// TIA Portal project "1215C_BREAKOUT_BOARD_IO-LINK_TEMPERATURE" (V19) (continued)
REGION Network 4: Add leading zero to HH:MM if less than 10
   // > If DTL.HOUR is less than 10 - replace 1st character in HH with a 0
   // > If DTL.MINUTE is less than 10 - replace 1st character in MM with a 0
   IF #LOCAL_DTL.HOUR < 10 THEN
       #sCustomTime_HH := REPLACE(IN1 := #sCustomTime_HH, IN2 := '0', L := 1, P := 1);
   END_IF;
   IF #LOCAL_DTL.MINUTE < 10 THEN
       #sCustomTime_MM := REPLACE(IN1 := #sCustomTime_MM, IN2 := '0', L := 1, P := 1);
   END_IF;
END_REGION

REGION Network 5: =================CONCAT_INTO_FORMAT=================
END_REGION

REGION Network 6: CONCAT Date into DD/MM/YY
   #sTemp_String := CONCAT(IN1 := #sCustomDate_DD, IN2 := '/');
   #sTemp_String := CONCAT(IN1 := #sTemp_String, IN2 := #sCustomDate_MM);
   #sTemp_String := CONCAT(IN1 := #sTemp_String, IN2 := '/');
   #sCustomDate_DDMMYY := CONCAT(IN1 := #sTemp_String, IN2 := #sCustomDate_YY);
END_REGION

REGION Network 7: CONCAT Time HH:MM
   #sCustomTime_HHMM := CONCAT(IN1 := #sCustomTime_HH, IN2 := ':');
   #sCustomTime_HHMM := CONCAT(IN1 := #sCustomTime_HHMM, IN2 := #sCustomTime_MM);
END_REGION
END_FUNCTION

// folder: WS01_TVET_Workstation/02-IOLink_Control

FUNCTION "FC10111-IFM_2Byte_PD" : Void   // FC10111, SCL
TITLE = IFM 2 Byte Process Data FC
{ S7_Optimized_Access := 'TRUE' }
VERSION : 0.1
// This function block is for a device with two byte process data input and no switch point in the 
// process data stream.
   VAR_INPUT
      I_PV : Int;   // input process value from master
      Gradient : Real;   // gradient see IODD descrption
   END_VAR
   VAR_OUTPUT
      O_PV_C : Real;   // output process value in deg c
      O_PV_F : Real;   // output process value in deg f
   END_VAR
   VAR_TEMP
      Temp_PV_C : Real;   // temp process value in deg c
   END_VAR
BEGIN
   // Convert input value using the gradient (default = 0.1)
   IF #Gradient > 0 THEN
       #Temp_PV_C := INT_TO_REAL(#I_PV) * #Gradient;
   ELSE
       #O_PV_C := INT_TO_REAL(#I_PV) * 1.0;
   END_IF;

   // Convert C to F
   #O_PV_F := (#Temp_PV_C * 1.8) + 32;

   // Move Temp_PV_C to O_PV_C
   #O_PV_C := #Temp_PV_C;
END_FUNCTION

// ===== library types =====

// folder: S7-1200/1500/Lib/S7-1200/1500/Common

FUNCTION_BLOCK "IO_LINK_DEVICE"   // FB50001, SCL
TITLE = IO_LINK_DEVICE
{ S7_Optimized_Access := 'TRUE' }
AUTHOR : SUP_FA
FAMILY : IO-Link
VERSION : 3.0
// Function block to read and write acyclic data on devices with IO-Link used on SIMATIC S7 controllers. (former IO_LINK_CALL)
   VAR_INPUT
      REQ : Bool;   // request function / Request Function / Neuer Auftrag
      ID : HW_IO;   // hardware identifier of IO-Link master module (HW_IO) from hw-config / Hardwarekennung des IOL-Master Moduls (HW_IO) aus HW-Konfiguration
      CAP : DInt := DINT#0;   // Client Access Point (CAP), for ET200 always 227 decimal / Client Access Point (CAP), bei ET200 immer 227 dez
      RD_WR : Bool;   // read and write access on IO-Link device 0: read, 1: write / Lese und Schreibzugriff auf IO-Link Device 0: Lesen, 1: schreiben
      PORT : Int := INT#0;   // number of port on IO-Link master module (ET200SP = 0..4) / Port/ Kanalnummer an dem das IO-Link Device betrieben wird. (ET200 = 0 .. 4)
      IOL_INDEX : Int := INT#0;   // address parameter Index (IO-Link Device) 0..32767 IOL-D, 65535 port functions / Adressparameter Index (IO-Link Device) 0..32767 IOL-D, 65535 port functions
      IOL_SUBINDEX : Int := INT#0;   // address parameter Subindex (IO-Link Device) 0 full record; 1-255 single parameter / Adressparameter Subindex (IO-Link Device) 0 ges. Record; 1-255 einz. Parameter
      LEN : Int := INT#0;   // length of writing data (netto data) / Länge der zu schreibenden Daten (Nettodaten)
   END_VAR
   VAR_OUTPUT
      DONE_VALID : Bool;   // validity 0: data invalid ; 1: data valid / Gültigkeit 0: Daten nicht gültig; 1: Daten gültig
      BUSY : Bool;   // 0: request finish 1: request in progress / 0: Auftrag abgeschlossen 1: Auftrag in Bearbeitung
      ERROR : Bool;   // Error Flag = 0: no error; 1: function aborted with error / Fehler Flag 0: kein Fehler; 1: Abbruch der Funktion mit Fehler
      STATUS : DWord := DW#16#00000000;   // DP/ PNIO - error status ; ERROR Flag = 1 - communication error status in detail / DP/ PNIO - Fehlerstatus; ERROR Flag = 1 - detaillierter Kommunikationsfehlerstatus
      IOL_STATUS : DWord := DW#16#00000000;   // IO-Link error status; ERROR flag = 1: IO-Link error status in detail / IO-Link Fehlerstatus; ERROR Flag = 1 - detaillierte IO-Link Fehlerstatus
      RD_LEN : Int := INT#0;   // length of read data record (number of bytes) / Länge des gelesenen Datensatzes (Anzahl Bytes)
   END_VAR
   VAR_IN_OUT
      RECORD_IOL_DATA : Array[0..231] of Byte;   // data area for reading / writing data (max. 232 byte) / Datenbereich für LESEN / SCHREIBEN (max. 232 Byte)
   END_VAR
   VAR
      RDREC_Function : RDREC;   // system function "read data record" (former SFB52) / Funktion Datensatz lesen (ehemals SFB52)
      WRREC_Function : WRREC;   // system function "write data record" (former SFB53) / Funktion Datensatz schreiben (ehemals SFB53)
      TP_poll : TP_TIME;   // poll rate read data record / Pollzeit für "Datensatz lesen"
      TON_monitoring : TON_TIME;   // request monitoring time / Überwachungszeit für Aufträge
      rdrec : Struct   // internal structure for RDREC / interne Struktur für RDREC
         valid : Bool;   // Function performed
         busy : Bool;   // Function busy
         error : Bool;   // Error flag
         status : DWord;   // Function result/error message
         length : UInt;   // Length of the fetched data record
      END_STRUCT;
      wrrec : Struct   // internal structure for WRREC / interne Struktur für WRREC
         length : UInt;   // length of write data record
         done : Bool;   // Function performed
         busy : Bool;   // Function busy
         error : Bool;   // Error flag
         status : DWord;   // Function result/error message
      END_STRUCT;
      read : Struct   // data area for reading data / Datenbereich für Lesedaten
         header : Struct
            CALL : Struct   // header for read/write data record
               Extended_Function_Num : Byte := 16#8;   // extended function number (fix coded 08h)
               Port : Byte;   // variable port (user interface) 0...255
               FI_Index : Word := 16#FE4A;   // FI index (fix coded 65098)
            END_STRUCT;
            IOL : Struct   // header for IO-Link
               Control : Byte;   // RD_WR = 0 = read = Control:=0x03 / / RD_WR = 1 = write = Control:=0x02
               Index_HighByte : Byte;   // index of data record 0…32767 (high byte)
               Index_LowByte : Byte;   // index of data record 0…32767 (low byte)
               Subindex : Byte;   // subindex for data record 0...255
            END_STRUCT;
         END_STRUCT;
         data : Array[0..231] of Byte;
      END_STRUCT;
      write : Struct   // data area for writing data / Datenbereich für Schreibdaten
         header : Struct
            CALL : Struct   // header for read/write data record
               Extended_Function_Num : Byte := 16#8;   // extended function number (fix coded 08h)
               Port : Byte;   // variable port (user interface) 0...255
               FI_Index : Word := 16#FE4A;   // FI index (fix coded 65098)
            END_STRUCT;
            IOL : Struct   // header for IO-Link
               Control : Byte;   // RD_WR = 0 = read = Control:=0x03 / / RD_WR = 1 = write = Control:=0x02
               Index_HighByte : Byte;   // index of data record 0…32767 (high byte)
               Index_LowByte : Byte;   // index of data record 0…32767 (low byte)
               Subindex : Byte;   // subindex for data record 0...255
            END_STRUCT;
         END_STRUCT;
         data : Array[0..231] of Byte;
      END_STRUCT;
      sequencecontrol : Int := INT#0;   // number of sequence control
      typeofrequest : Int := INT#0;   // type of request (0=Read, 1=Write)
      R_TRIG_REQ : Bool;   // impulse start new request / Impuls für neuen Auftrag starten
      R_TRIG_REQ_old : Bool;   // old value of REQ (previous cycle) / Flankenmerker
      F_TRIG_poll : Bool;   // impulse poll read data record (response) / Impuls für Pollen "Datensatz lesen"
      F_TRIG_poll_old : Bool;   // old value of Poll (previous cycle) / Flankenmerker
   END_VAR
   VAR_TEMP
      retval : Int;   // function return value / Variable für Rückgabewerte von Funktionen
      tmpWORD : Word;   // data type WORD for temporarily use / Datentyp WORD zur temporären Verwendung
      tmpDWORD : DWord;   // data type DWORD for temporarily use / Datentyp DWORD zur temporären Verwendung
      tmpINT : Int;   // data type INT for temporarily use / Datentyp INT zur temporären Verwendung
      i : Int;   // run tag for counting loops / Laufvariable für for-Schleifen
   END_VAR
BEGIN
   (*---------------------------------------------------------------------------------------------------------------------
   SIEMENS AG
   ©Copyright 2015. All Rights Reserved.
   -----------------------------------------------------------------------------------------------------------------------
   Limitation of liability
   This software was developed with largest care. However, the author can not guarantee, that the software runs under
   each version of STEP7 on each PLC flawlessly.
   There is no warranty for the software, to the extent permitted by applicable law. The copyright holder provides the
   software "as is" without warranty of any kind, either expressed or implied, including, but not limited to, the implied
   warranties of merchantability and fitness for a particular purpose. The entire risk as to the quality and performance
   of the software is with you. Should the software prove defective, you assume the cost of all necessary servicing,
   repair or correction. In no event unless required by applicable law will the copyright holder be liable to you for
   damages, including any general, special, incidental or consequential damages arising out of the use or inability to
   use the software (including but not limited to loss of data or data being rendered inaccurate or losses sustained by
   you or third parties or a failure of the software to operate with any other programs), even if such holder or other
   party has been advised of the possibility of such damages.
   Permission to use or copy this software for any purpose is hereby granted without fee, provided the above notices are
   retained on all copies. Permission to modify the code and to distribute modified code is granted, provided the above
   notices are retained, and a notice that the code was modified is included with the above copyright notice.
   -----------------------------------------------------------------------------------------------------------------------
   Functionality provided by this source (short description):
   Function block IO_LINK_DEVICE - used to read and write of acyclic data records on devices with IO-Link.
   Note:
   To read data records, the IO-Link master modules needs to know which data record is required. Therefore it is necessary
   to send at first a request via write data record (only header of 8 byte). As response the IO-Link master module
   will send the required data record.

   Status:     Released (tested)
   File name:  IO_LINK_DEVICE
   System :    SIMATIC S7-1200/1500
   Version :   3.0
   -----------------------------------------------------------------------------------------------------------------------
   Script to be stored on level ... in project (mark appropriate levels with [x] below)
   [ ] External
   [ ] All levels possible
   [x] Project level
   [ ] Controller level
   [ ] Device level
   [ ] Subobject level
   -----------------------------------------------------------------------------------------------------------------------
   Restrictions, known limitations:
   The limitation of 240 byte is based on PROFIBUS DP protocol. With PROFINET IO there wouldn't no limit but because of 
   compatibility reason it wasn't changed.
     - header =   8 byte
     - data   = 232 byte
   -----------------------------------------------------------------------------------------------------------------------
   Requirements, prerequisites, External resources used: nothing
   -----------------------------------------------------------------------------------------------------------------------
   Change log table (latest change is at the bottom OF the list):
   Version Date Changes applied
   V2.0.0 <2013-09-30> First created with TIA Portal V12 SP1
   V2.1.0 <2014-03-14> Upgrade system function 'WRREC' from V1.0 to V1.1 and released for TIA Portal V13
   V3.0.0 <2015-02-28> Upgrade and released for TIA Portal V13 SP1 (without backup/restore master parameter)
   V3.0.2 <2015-07-07> Change of #IOL_INDEX and #Port lower boundry to 0
   ---------------------------------------------------------------------------------------------------------------------*)

   (*---------------------------------------------------------------------------------------------------------------------
   Description of programmed IO-Link error codes
   8000 = time out
   8001 = wrong port
   8002 = wrong index
   8003 = wrong subindex
   8005 = wrong length for write data record
   8006 = wrong length for read data record
   8052 = error during reading data record
   8053 = error during writing data record
   All other codes are coming from a higher level!
   ---------------------------------------------------------------------------------------------------------------------*)

   (*---------------------------------------------------------------------------------------------------------------------
               NEW REQUEST
   ---------------------------------------------------------------------------------------------------------------------*)
   // detection rising edge of "REQ"
   #R_TRIG_REQ := #REQ = TRUE AND #R_TRIG_REQ_old = FALSE;
   #R_TRIG_REQ_old := #REQ = TRUE;

   // start new request if not busy
   IF #R_TRIG_REQ = TRUE AND #sequencecontrol = 0 THEN
       // Freeze record ID and CAP
       #WRREC_Function.ID := #ID;
       #WRREC_Function.INDEX := #CAP;
       #RDREC_Function.ID := #ID;
       #RDREC_Function.INDEX := #CAP;

       // Initialize outputs
       #DONE_VALID := FALSE;
       #BUSY := TRUE;
       #ERROR := FALSE;
       #STATUS := DW#16#00000000;
       #IOL_STATUS := DW#16#00000000;
       #RD_LEN := INT#0;

       // Initialize data area
       #read.header.CALL.Port := B#16#0;
       #read.header.IOL.Index_LowByte := B#16#0;
       #read.header.IOL.Index_HighByte := B#16#0;
       #read.header.IOL.Subindex := B#16#0;
       #i := INT#0; // initialize loop counter      
       FOR #i := 0 TO 231 DO
           #write.data[#i] := B#16#0;
           #read.data[#i] := B#16#0;
       END_FOR;

   (*---------------------------------------------------------------------------------------------------------------------
       Setup IO-LINK Call needs a specific header
   ---------------------------------------------------------------------------------------------------------------------*)
   // setup CALL header
   #write.header.CALL.Extended_Function_Num := 16#08;  // extended function number (fix coded 08h)
   #write.header.CALL.Port := INT_TO_BYTE(#PORT);  // 1..63 = PORT number, 64..255=reserved
   #write.header.CALL.FI_Index := 65098;  // IOL-Header is following (fix coded 65098)

   // setup IOL header 
   // CONTROL = please see below at BODY
   // INDEX
   #write.header.IOL.Index_LowByte := INT_TO_BYTE(#IOL_INDEX);
   #tmpWORD := INT_TO_WORD(#IOL_INDEX);
   #tmpWORD := SHR(IN := #tmpWORD, N := 8);
   #write.header.IOL.Index_HighByte := WORD_TO_BYTE(#tmpWORD);
   // SUBINDEX
   #write.header.IOL.Subindex := INT_TO_BYTE(#IOL_SUBINDEX);

   // BODY (data max. 232 Byte, Array 0..231 of Byte) 
   IF #RD_WR = TRUE THEN
       // IO-Link write data record requested, copy data from "RECORD_IOL_DATA"
       #write.header.IOL.Control := B#16#02; // CONTROL B#16#02 = write data record
       #wrrec.length := INT_TO_UINT(#LEN) + UINT#8;  // data length header + data = IO-Link write data record
       #typeofrequest := 2; // write data record
       // copy IOL_RECORD_DATA in working area
       #i := INT#0;    // initialize loop counter 
       FOR #i := 0 TO #LEN - 1 DO
           #write.data[#i] := #RECORD_IOL_DATA[#i];
       END_FOR;
   ELSE
       // IO-Link read data record requested
       #write.header.IOL.Control := 16#03;  // CONTROL 16#03 = read data record
       #wrrec.length := UINT#8; // data length only header = IO-Link read data record
       #typeofrequest := 1; // read data record        
   END_IF;
   #sequencecontrol := 1;  // Start sequence
   ELSE
       ;
   END_IF;

   (*---------------------------------------------------------------------------------------------------------------------
               SEQUENCE CONTROL
   ---------------------------------------------------------------------------------------------------------------------*)
   CASE #sequencecontrol OF
       1:  // Check input parameter        
           IF #PORT < INT#0 OR #PORT > INT#63 THEN // PORT (Wrong port address = 0x8001)
               #ERROR := TRUE;
               #IOL_STATUS := DW#16#80010000;
               #sequencecontrol := 99; // aborting function with error
           ELSIF #IOL_INDEX < INT#0 OR #IOL_INDEX > INT#32767 THEN    // INDEX (Wrong index = 0x8002)
               #ERROR := TRUE;
               #IOL_STATUS := DW#16#80020000;
               #sequencecontrol := 99; // aborting function with error
           ELSIF #IOL_SUBINDEX < INT#0 OR #IOL_SUBINDEX > INT#255 THEN    // SUBINDEX (Wrong subindex = 0x8003)
               #ERROR := TRUE;
               #IOL_STATUS := DW#16#80030000;
               #sequencecontrol := 99; // aborting function with error
           ELSIF #typeofrequest = 2 AND (#LEN < 1 OR #LEN > 232) THEN  // LEN (wrong length for write data record = 0x8004)
               #ERROR := TRUE;
               #IOL_STATUS := DW#16#80050000;
               #sequencecontrol := 99; // aborting function with error
           ELSIF #typeofrequest = 1 AND (#LEN < 0 OR #LEN > 232) THEN  // LEN (wrong length for read data record = 0x8005)
               #ERROR := TRUE;
               #IOL_STATUS := DW#16#80060000;
               #sequencecontrol := 99; // aborting function with error
           ELSE    // all input parameter are right
               #sequencecontrol := 2;
           END_IF;

       2:  (*-------------------------------------------------------------------------------------------------------------
           WRREC = Write Data Record
           Note:
           To read data records, the IO-Link master modules needs to know which PORT is required. Therefore it is necessary
           to send at first a request via write data record (header, 8 byte). As response the IO-Link master module will 
           send the required data record.
           -------------------------------------------------------------------------------------------------------------*)
           #WRREC_Function(REQ := TRUE,
                           LEN := #wrrec.length,
                           DONE => #wrrec.done,
                           BUSY => #wrrec.busy,
                           ERROR => #wrrec.error,
                           STATUS => #wrrec.status,
                           RECORD := #write);
           // output status during write data record
           IF #wrrec.busy THEN
               #STATUS := #wrrec.status;
               #IOL_STATUS := DW#16#00020000;  // 0002 = writing in progress 
           ELSIF #wrrec.error THEN
               #tmpDWORD := #wrrec.status AND DW#16#00FFFF00;  // filter status
               IF #tmpDWORD = DW#16#0080C200 THEN    // if resource #BUSY (#STATUS=80C2), then ... 
                   #sequencecontrol := 3;  // ... repeat write data record
               ELSE
                   #ERROR := TRUE;
                   #STATUS := #wrrec.status;   // ... otherwise output error status of "WRREC"
                   #IOL_STATUS := DW#16#80530000;  // ... with note '8053' = error status of "WRREC"
                   #sequencecontrol := 99; // aborting function with error
               END_IF;
           ELSIF #wrrec.done = TRUE THEN   // wait for write data record finish without error
               #TP_poll(IN := TRUE,
                        PT := T#100ms);    // poll for response
               #sequencecontrol := 4;
           ELSE
               ;
           END_IF;

       3:  // repeat write data record because resource was busy
           #WRREC_Function(REQ := FALSE);
           #sequencecontrol := 2;

       4:  // wait and poll for response = Read Data Record (RDREC)
           #WRREC_Function(REQ := FALSE);
           #TP_poll(IN := TRUE,
                    PT := T#100ms);

           // if poll rate executed then start read data record (on falling edge)
           #F_TRIG_poll := #TP_poll.Q = FALSE AND #F_TRIG_poll_old = TRUE;
           #F_TRIG_poll_old := #TP_poll.Q = TRUE;

           // RDREC = Read Data Record
           #RDREC_Function(REQ := #F_TRIG_poll,
                           MLEN := UINT#0, // length = 0 = read all data which are available
                           VALID => #rdrec.valid,
                           BUSY => #rdrec.busy,
                           ERROR => #rdrec.error,
                           STATUS => #rdrec.status,
                           LEN => #rdrec.length,
                           RECORD := #read);
           // output status during read data record
           IF #rdrec.busy THEN
               #STATUS := #rdrec.status;
               #IOL_STATUS := DW#16#00030000; // 16#0003 = reading in progress
           ELSIF #rdrec.error = TRUE THEN
               #tmpDWORD := #rdrec.status AND DW#16#00FFFF00;  // filter status
               IF #tmpDWORD = DW#16#0080C200 THEN  // if resource busy (status=80C2), then ... 
                   #sequencecontrol := 5;  // ... repeat read data record / continue polling
               ELSE
                   #ERROR := TRUE;
                   #STATUS := #rdrec.status;   // ... otherwise output error code of "RDREC"
                   #IOL_STATUS := DW#16#80520000;  // ... with note '8052' = error status of "RDREC"
                   #sequencecontrol := 99; // aborting function with error
               END_IF;
           ELSIF #rdrec.valid THEN
               IF  // check the response wether it matches the request (compare PORT, INDEX and SUBINDEX)
                   (#write.header.CALL.Port <> #read.header.CALL.Port) OR
                   (#write.header.IOL.Index_HighByte <> #read.header.IOL.Index_HighByte) OR
                   (#write.header.IOL.Index_LowByte <> #read.header.IOL.Index_LowByte) OR
                   (#write.header.IOL.Subindex <> #read.header.IOL.Subindex)
               THEN    // read data record don't match the request
                   #ERROR := TRUE;
                   #STATUS := #rdrec.status;
                   #IOL_STATUS := DW#16#70000000;  // output status '7000', no consistent data
                   #sequencecontrol := 99; // aborting function with error
               ELSIF #read.header.IOL.Control = B#16#80 THEN   // check the response for IO-Link errors
                   // State 0x80 = IOL_CALL_RES PDU shows IO-Link error detect
                   #ERROR := TRUE;
                   #STATUS := DW#16#00000000;
                   #IOL_STATUS.%B3 := #read.data[0];   // IO-Link master error code
                   #IOL_STATUS.%B2 := #read.data[1];   // IO-Link master error code
                   #IOL_STATUS.%B1 := #read.data[2];  // IO-Link device error code
                   #IOL_STATUS.%B0 := #read.data[3];  // IO-Link device additional error code

                   #sequencecontrol := 99; // aborting function with error
               ELSE    // read data are valid = output
                   #DONE_VALID := TRUE;
                   #BUSY := FALSE;
                   #ERROR := FALSE;
                   #STATUS := DW#16#00000000;
                   #IOL_STATUS := DW#16#00000000;  // request finished

                   IF #typeofrequest = 1 THEN
                       #RD_LEN := UINT_TO_INT(#rdrec.length - UINT#8);  // device parameter cover header and data,
                       // only data will be output
                       #i := INT#0; // initialize loop counter
                       FOR #i := 0 TO UINT_TO_INT(#rdrec.length - UINT#8 - UINT#1) DO
                           #RECORD_IOL_DATA[#i] := #read.data[#i];
                       END_FOR;
                   ELSE
                       ;
                   END_IF;
                   #sequencecontrol := 98;
               END_IF;
           ELSE
               ;
           END_IF;

       5:  // poll again for response because resource was busy
           #TP_poll(IN := FALSE,
                    PT := T#100ms);
           #RDREC_Function(REQ := FALSE,
                           RECORD := #read);
           #sequencecontrol := 4;  // ... repeat read data record / continue polling   

       98: // request done successfully
           #TP_poll(IN := FALSE,
                    PT := T#100ms);
           #RDREC_Function(REQ := FALSE,
                           RECORD := #read);
           IF #REQ = FALSE THEN
               #DONE_VALID := FALSE;
               #BUSY := FALSE;
               #ERROR := FALSE;
               #RD_LEN := INT#0;
               #STATUS := DW#16#00000000;
               #IOL_STATUS := DW#16#00010000; // ready for new request
               #sequencecontrol := 0;
               #typeofrequest := 0;
           ELSE
               ;
           END_IF;

       99: // Function aborted with error
           #TP_poll(IN := FALSE,
                    PT := T#100ms);
           #WRREC_Function(REQ := FALSE);
           #RDREC_Function(REQ := FALSE,
                           RECORD := #read);
           #DONE_VALID := FALSE;
           #BUSY := FALSE;
           #RD_LEN := INT#0;
           #sequencecontrol := 0;
           #typeofrequest := 0;

       ELSE  // no relevant case, ready for new request
           #WRREC_Function(REQ := FALSE);
           #RDREC_Function(REQ := FALSE,
                           RECORD := #read);
           #TP_poll(IN := FALSE,
                    PT := T#100ms);
           #TON_monitoring(IN := FALSE,
                           PT := T#20s);
           #sequencecontrol := 0;
           #typeofrequest := 0;
   END_CASE;

   (*---------------------------------------------------------------------------------------------------------------------
               MONITORING
   ---------------------------------------------------------------------------------------------------------------------*)
   #TON_monitoring(IN := #sequencecontrol > 0 AND #sequencecontrol < 98,
                   PT := T#20s);
   IF #TON_monitoring.Q THEN
       #ERROR := TRUE;
       #IOL_STATUS := DW#16#80000000; // request time out       
       #sequencecontrol := 99; // aborting function with error
   END_IF;
END_FUNCTION_BLOCK

(* ===== HMI "HMI_RT_1" =====
system functions are stored by id; their names below are inferred from use
connection "HMI_Connection": ETHERNET, SMART_S7_1200_OMS

HMI tags "Default tag table"
   "ScreenNumber" : UInt, internal

HMI tags "PLC_Inputs"
   "DB001-PLC_I/O_Inputs_xDI0.0" : Bool = PLC "DB001-PLC_I/O".Inputs."xDI0.0", 100 ms
   "DB001-PLC_I/O_Inputs_xDI0.1" : Bool = PLC "DB001-PLC_I/O".Inputs."xDI0.1", 100 ms
   "DB001-PLC_I/O_Inputs_xDI0.2" : Bool = PLC "DB001-PLC_I/O".Inputs."xDI0.2", 100 ms
   "DB001-PLC_I/O_Inputs_xDI0.3" : Bool = PLC "DB001-PLC_I/O".Inputs."xDI0.3", 100 ms
   "DB001-PLC_I/O_Inputs_xDI0.4" : Bool = PLC "DB001-PLC_I/O".Inputs."xDI0.4", 100 ms
   "DB001-PLC_I/O_Inputs_xDI0.5" : Bool = PLC "DB001-PLC_I/O".Inputs."xDI0.5", 100 ms
   "DB001-PLC_I/O_Inputs_xDI0.6" : Bool = PLC "DB001-PLC_I/O".Inputs."xDI0.6", 100 ms
   "DB001-PLC_I/O_Inputs_xDI0.7" : Bool = PLC "DB001-PLC_I/O".Inputs."xDI0.7", 100 ms
   "DB001-PLC_I/O_Inputs_xDI1.0" : Bool = PLC "DB001-PLC_I/O".Inputs."xDI1.0", 100 ms
   "DB001-PLC_I/O_Inputs_xDI1.1" : Bool = PLC "DB001-PLC_I/O".Inputs."xDI1.1", 100 ms
   "DB001-PLC_I/O_Inputs_xDI1.2" : Bool = PLC "DB001-PLC_I/O".Inputs."xDI1.2", 100 ms
   "DB001-PLC_I/O_Inputs_xDI1.3" : Bool = PLC "DB001-PLC_I/O".Inputs."xDI1.3", 100 ms
   "DB001-PLC_I/O_Inputs_xDI1.4" : Bool = PLC "DB001-PLC_I/O".Inputs."xDI1.4", 100 ms
   "DB001-PLC_I/O_Inputs_xDI1.5" : Bool = PLC "DB001-PLC_I/O".Inputs."xDI1.5", 100 ms

HMI tags "PLC_Outputs"
   "DB001-PLC_I/O_Outputs_xDQ0.0" : Bool = PLC "DB001-PLC_I/O".Outputs."xDQ0.0", 100 ms
   "DB001-PLC_I/O_Outputs_xDQ0.1" : Bool = PLC "DB001-PLC_I/O".Outputs."xDQ0.1", 100 ms
   "DB001-PLC_I/O_Outputs_xDQ0.2" : Bool = PLC "DB001-PLC_I/O".Outputs."xDQ0.2", 100 ms
   "DB001-PLC_I/O_Outputs_xDQ0.3" : Bool = PLC "DB001-PLC_I/O".Outputs."xDQ0.3", 100 ms
   "DB001-PLC_I/O_Outputs_xDQ0.4" : Bool = PLC "DB001-PLC_I/O".Outputs."xDQ0.4", 100 ms
   "DB001-PLC_I/O_Outputs_xDQ0.5" : Bool = PLC "DB001-PLC_I/O".Outputs."xDQ0.5", 100 ms
   "DB001-PLC_I/O_Outputs_xDQ0.6" : Bool = PLC "DB001-PLC_I/O".Outputs."xDQ0.6", 100 ms
   "DB001-PLC_I/O_Outputs_xDQ0.7" : Bool = PLC "DB001-PLC_I/O".Outputs."xDQ0.7", 100 ms
   "DB001-PLC_I/O_Outputs_xDQ1.0" : Bool = PLC "DB001-PLC_I/O".Outputs."xDQ1.0", 100 ms
   "DB001-PLC_I/O_Outputs_xDQ1.1" : Bool = PLC "DB001-PLC_I/O".Outputs."xDQ1.1", 100 ms

HMI tags "PLC_Analog"
   "AI0.0" : Word = PLC "AI0.0" AT %IW64, 100 ms
   "AQ0.0" : Word = PLC "AQ0.0" AT %QW64, 100 ms
   "DB001-PLC_I/O_Outputs_rAQ0.0_Scaled" : Real = PLC "DB001-PLC_I/O".Inputs."rAI0.0_Scaled", 100 ms
   "DB001-PLC_I/O_Outputs_rAQ0.1_Scaled" : Real = PLC "DB001-PLC_I/O".Inputs."rAI0.1_Scaled", 100 ms
   "AI0.1" : Word = PLC "AI0.1" AT %IW66, 100 ms
   "AQ0.1" : Word = PLC "AQ0.1" AT %QW66, 100 ms
   "DB001-PLC_I/O_Inputs_rAI0.0_Scaled" : Real = PLC "DB001-PLC_I/O".Inputs."rAI0.0_Scaled", 100 ms
   "DB001-PLC_I/O_Inputs_rAI0.1_Scaled" : Real = PLC "DB001-PLC_I/O".Inputs."rAI0.1_Scaled", 100 ms

HMI tags "PLC_DateTime"
   "DB002-DateTime_sCustomDate_DDMMYY" : String[254] = PLC "DB002-DateTime".sCustomDate_DDMMYY, 100 ms
   "DB002-DateTime_sCustomTime_HHMM" : String[254] = PLC "DB002-DateTime".sCustomTime_HHMM, 100 ms

HMI tags "IO-Link"
   "DB003-IOLink_Data_TempSensor_Data_rDeg_C" : Real = PLC "DB004-IOLink_Data".TempSensor_Data.rDeg_C, 100 ms
   "DB003-IOLink_Data_TempSensor_Data_rDeg_F" : Real = PLC "DB004-IOLink_Data".TempSensor_Data.rDeg_F, 100 ms

text list "ON/OFF": 0 'OFF'; 1 'ON'

screen "01-Home" 480x272, template "Main_Template"
   on GenerateScreen: SetTag("ScreenNumber", 1)
   TextField "TextField_ProjectName" at 109,47 size 259x30; Text 'PLC BREAKOUT BOARD'
   TextField "Text field_DeviceInfo" at 21,85 size 435x52; Text '1215C DC/DC/DC -- 6ES7215-1AG40-0XB0 -- IP: 192.168.0.175/24 KTP400 HMI -- 6AV2123-2DB03-0AX0 -- IP: 192.168.0.176/24 IFM IO-LINK MASTER -- AL1100 -- IP: 192.168.0.177/24'
   TextField "Text field_Description" at 62,143 size 353x68; Text '- Displays the Digital & Analog Input states, - Toggle Digital Outputs via HMI buttons, - Simulation of Analog Outputs via 20 step incriments, - Manipulation of the IO-Link temperature reading.'
   Button "Button_ExitRuntime" at 384,227 size 92x40; TextOff 'EXIT RUNTIME'
      on Press: StopRuntime(0)

screen "02-Inputs1" 480x272, template "Main_Template"
   on GenerateScreen: SetTag("ScreenNumber", 2)
   TextField "TextField_ScreenName" at 85,46 size 309x30; Text 'PLC DIGITAL INPUTS - 1of3'
   TextField "TextField_BankLetter" at 412,50 size 64x23; Text 'BANK A'
   Button "Button_Next" at 384,227 size 92x40; TextOff 'NEXT'
      on Press: ActivateScreen("03-Inputs2", 0)
   Group "Group_DI0.0" at 41,81 size 62x63
   Group "Group_DI0.1" at 153,81 size 62x63
   Group "Group_DI0.2" at 265,81 size 62x63
   Group "Group_DI0.3" at 377,81 size 62x63
   Group "Group_DI0.4" at 41,152 size 62x64
   Group "Group_DI0.5" at 153,152 size 62x64
   Group "Group_DI0.6" at 265,154 size 62x64
   Group "Group_DI0.7" at 377,154 size 62x64
   TextField "Text field_DI0.0" at 51,81 size 42x19; Text 'DI 0.0'
   Circle "Circle_DI0.0" at 54,103 size 36x36
      Appearance <- "DB001-PLC_I/O_Inputs_xDI0.0"
   TextField "Text field_DI0.1" at 163,81 size 42x19; Text 'DI 0.1'
   Circle "Circle_DI0.1" at 166,103 size 36x36
      Appearance <- "DB001-PLC_I/O_Inputs_xDI0.1"
   TextField "Text field_DI0.2" at 275,81 size 42x19; Text 'DI 0.2'
   Circle "Circle_DI0.2" at 278,103 size 36x36
      Appearance <- "DB001-PLC_I/O_Inputs_xDI0.2"
   TextField "Text field_DI0.3" at 387,81 size 42x19; Text 'DI 0.3'
   Circle "Circle_DI0.3" at 390,103 size 36x36
      Appearance <- "DB001-PLC_I/O_Inputs_xDI0.3"
   TextField "Text field_DI0.4" at 51,152 size 42x19; Text 'DI 0.4'
   Circle "Circle_DI0.4" at 54,174 size 36x36
      Appearance <- "DB001-PLC_I/O_Inputs_xDI0.4"
   TextField "Text field_DI0.5" at 163,152 size 42x19; Text 'DI 0.5'
   Circle "Circle_DI0.5" at 166,174 size 36x36
      Appearance <- "DB001-PLC_I/O_Inputs_xDI0.5"
   TextField "Text field_DI0.6" at 275,154 size 42x19; Text 'DI 0.6'
   Circle "Circle_DI0.6" at 278,176 size 36x36
      Appearance <- "DB001-PLC_I/O_Inputs_xDI0.6"
   TextField "Text field_DI0.7" at 387,154 size 42x19; Text 'DI 0.7'
   Circle "Circle_DI0.7" at 390,176 size 36x36
      Appearance <- "DB001-PLC_I/O_Inputs_xDI0.7"

screen "05-Outputs1" 480x272, template "Main_Template"
   on GenerateScreen: SetTag("ScreenNumber", 5)
   TextField "TextField_ScreenName" at 76,46 size 328x30; Text 'PLC DIGITAL OUTPUTS - 1of3'
   TextField "TextField_BankLetter" at 412,50 size 64x23; Text 'BANK A'
   Button "Button_Next" at 384,227 size 92x40; TextOff 'NEXT'
      on Press: ActivateScreen("06-Outputs2", 0)
   Group "Group_DQ0.0" at 18,83 size 97x62; TextList "ON/OFF"
   Group "Group_DQ0.1" at 132,83 size 97x62; TextList "ON/OFF"
   Group "Group_DQ0.2" at 247,83 size 97x62; TextList "ON/OFF"
   Group "Group_DQ0.3" at 362,83 size 97x62; TextList "ON/OFF"
   Group "Group_DQ0.4" at 18,154 size 97x62; TextList "ON/OFF"
   Group "Group_DQ0.5" at 132,154 size 97x62; TextList "ON/OFF"
   Group "Group_DQ0.6" at 247,154 size 97x62; TextList "ON/OFF"
   Group "Group_DQ0.7" at 362,154 size 97x62; TextList "ON/OFF"
   Rectangle "Rectangle_DQ0.0" at 18,83 size 97x62
      Appearance <- "DB001-PLC_I/O_Outputs_xDQ0.0"
   TextField "Text field_DQ0.0" at 44,83 size 46x19; Text 'DQ 0.0'
   Button "Button_DQ0.0" at 30,105 size 73x32; TextOff 'Text'; TextList "ON/OFF"
      on Press: InvertBit("DB001-PLC_I/O_Outputs_xDQ0.0")
      ProcessValue <- "DB001-PLC_I/O_Outputs_xDQ0.0"
   Rectangle "Rectangle_DQ0.1" at 132,83 size 97x62
      Appearance <- "DB001-PLC_I/O_Outputs_xDQ0.1"
   TextField "Text field_DQ0.1" at 158,83 size 46x19; Text 'DQ 0.1'
   Button "Button_DQ0.1" at 144,105 size 73x32; TextOff 'Text'; TextList "ON/OFF"
      on Press: InvertBit("DB001-PLC_I/O_Outputs_xDQ0.1")
      ProcessValue <- "DB001-PLC_I/O_Outputs_xDQ0.1"
   Rectangle "Rectangle_DQ0.2" at 247,83 size 97x62
      Appearance <- "DB001-PLC_I/O_Outputs_xDQ0.2"
   TextField "Text field_DQ0.2" at 273,83 size 46x19; Text 'DQ 0.2'
   Button "Button_DQ0.2" at 259,105 size 73x32; TextOff 'Text'; TextList "ON/OFF"
      on Press: InvertBit("DB001-PLC_I/O_Outputs_xDQ0.2")
      ProcessValue <- "DB001-PLC_I/O_Outputs_xDQ0.2"
   Rectangle "Rectangle_DQ0.3" at 362,83 size 97x62
      Appearance <- "DB001-PLC_I/O_Outputs_xDQ0.3"
   TextField "Text field_DQ0.3" at 388,83 size 46x19; Text 'DQ 0.3'
   Button "Button_DQ0.3" at 374,105 size 73x32; TextOff 'Text'; TextList "ON/OFF"
      on Press: InvertBit("DB001-PLC_I/O_Outputs_xDQ0.3")
      ProcessValue <- "DB001-PLC_I/O_Outputs_xDQ0.3"
   Rectangle "Rectangle_DQ0.4" at 18,154 size 97x62
      Appearance <- "DB001-PLC_I/O_Outputs_xDQ0.4"
   TextField "Text field_DQ0.4" at 44,154 size 46x19; Text 'DQ 0.4'
   Button "Button_DQ0.4" at 30,176 size 73x32; TextOff 'Text'; TextList "ON/OFF"
      on Press: InvertBit("DB001-PLC_I/O_Outputs_xDQ0.4")
      ProcessValue <- "DB001-PLC_I/O_Outputs_xDQ0.4"
   Rectangle "Rectangle_DQ0.5" at 132,154 size 97x62
      Appearance <- "DB001-PLC_I/O_Outputs_xDQ0.5"
   TextField "Text field_DQ0.5" at 158,154 size 46x19; Text 'DQ 0.5'
   Button "Button_DQ0.5" at 144,176 size 73x32; TextOff 'Text'; TextList "ON/OFF"
      on Press: InvertBit("DB001-PLC_I/O_Outputs_xDQ0.5")
      ProcessValue <- "DB001-PLC_I/O_Outputs_xDQ0.5"
   Rectangle "Rectangle_DQ0.6" at 247,154 size 97x62
      Appearance <- "DB001-PLC_I/O_Outputs_xDQ0.6"
   TextField "Text field_DQ0.6" at 273,154 size 46x19; Text 'DQ 0.6'
   Button "Button_DQ0.6" at 259,176 size 73x32; TextOff 'Text'; TextList "ON/OFF"
      on Press: InvertBit("DB001-PLC_I/O_Outputs_xDQ0.6")
      ProcessValue <- "DB001-PLC_I/O_Outputs_xDQ0.6"
   Rectangle "Rectangle_DQ0.7" at 362,154 size 97x62
      Appearance <- "DB001-PLC_I/O_Outputs_xDQ0.7"
   TextField "Text field_DQ0.7" at 388,154 size 46x19; Text 'DQ 0.7'
   Button "Button_DQ0.7" at 374,176 size 73x32; TextOff 'Text'; TextList "ON/OFF"
      on Press: InvertBit("DB001-PLC_I/O_Outputs_xDQ0.7")
      ProcessValue <- "DB001-PLC_I/O_Outputs_xDQ0.7"

screen "08-AnalogI/O" 480x272, template "Main_Template"
   on GenerateScreen: SetTag("ScreenNumber", 8)
   Button "Button_Back" at 384,227 size 92x40; TextOff 'BACK'
      on Press: function_efd93a16()
   TextField "TextField_ScreenName" at 65,46 size 351x30; Text 'PLC ANALOG INPUTS/OUTPUTS'
   Group "Group_A0" at 244,76 size 229x145; FormatPattern 9999
   Group "Group_A1" at 8,76 size 229x145; FormatPattern 9999
   TextField "Text field_A0" at 291,77 size 127x21; Text 'Analog AI-0 & AQ-0'
   TextField "Text field_A0_Input" at 279,98 size 42x17; Text 'INPUT'
   TextField "Text field_A0_Instruction" at 256,115 size 86x34; Text 'Use the connected potentiometer to change the input voltage.'
   TextField "Text field_A0_Voltage" at 280,149 size 41x14; Text 'VOLTAGE:'
   IOField "I/O field_A0_Voltage" at 281,162 size 42x21; FormatPattern 99.99; Unit  V
      ProcessValue <- "DB001-PLC_I/O_Inputs_rAI0.0_Scaled"
   TextField "Text field_A0_InRAW" at 289,181 size 24x14; Text 'RAW:'
   IOField "I/O field_A0_RAW" at 283,193 size 37x21; FormatPattern 99999
      ProcessValue <- "AI0.0"
   TextField "Text field_A0_Output" at 389,98 size 52x17; Text 'OUTPUT'
   TextField "Text field_A0_mA" at 381,127 size 19x14; Text 'mA:'
   IOField "I/O field_A0_mA" at 365,140 size 51x21; FormatPattern 99.99; Unit  mA
      ProcessValue <- "DB001-PLC_I/O_Outputs_rAQ0.0_Scaled"
   TextField "Text field_A0_OutRAW" at 379,167 size 24x14; Text 'RAW:'
   IOField "I/O field_A0_OutRAW" at 373,180 size 37x21; FormatPattern 99999
      ProcessValue <- "AQ0.0"
   TextField "Text field_A0_20" at 403,113 size 25x14; Text '20mA'
   TextField "Text field_A0_15" at 415,136 size 13x14; Text '15'
   TextField "Text field_A0_10" at 415,160 size 13x14; Text '10'
   TextField "Text field_A0_5" at 419,182 size 10x14; Text '5'
   TextField "Text field_A0_0" at 408,205 size 21x14; Text '0mA'
   Bar "Bar_A0" at 428,118 size 37x97; MinimumValue 0; MaximumValue 20
      ProcessValue <- "DB001-PLC_I/O_Outputs_rAQ0.0_Scaled"
   TextField "Text field_A1" at 55,77 size 127x21; Text 'Analog AI-1 & AQ-1'
   TextField "Text field_A1_Input" at 43,98 size 42x17; Text 'INPUT'
   TextField "Text field_A1_Instruction" at 20,115 size 86x34; Text 'Use the connected potentiometer to change the input voltage.'
   TextField "Text field_A1_Voltage" at 44,149 size 41x14; Text 'VOLTAGE:'
   IOField "I/O field_A1_Voltage" at 45,162 size 42x21; FormatPattern 99.99; Unit  V
      ProcessValue <- "DB001-PLC_I/O_Inputs_rAI0.1_Scaled"
   TextField "Text field_A1_InRAW" at 53,181 size 24x14; Text 'RAW:'
   IOField "I/O field_A1_RAW" at 47,193 size 37x21; FormatPattern 99999
      ProcessValue <- "AI0.1"
   TextField "Text field_A1_Output" at 153,98 size 52x17; Text 'OUTPUT'
   TextField "Text field_A1_mA" at 145,127 size 19x14; Text 'mA:'
   IOField "I/O field_A1_mA" at 129,140 size 51x21; FormatPattern 99.99; Unit  mA
      ProcessValue <- "DB001-PLC_I/O_Outputs_rAQ0.1_Scaled"
   TextField "Text field_A1_OutRAW" at 143,167 size 24x14; Text 'RAW:'
   IOField "I/O field_A1_OutRAW" at 137,180 size 37x21; FormatPattern 99999
      ProcessValue <- "AQ0.1"
   TextField "Text field_A1_20" at 167,113 size 25x14; Text '20mA'
   TextField "Text field_A1_15" at 179,136 size 13x14; Text '15'
   TextField "Text field_A1_10" at 179,160 size 13x14; Text '10'
   TextField "Text field_A1_5" at 183,182 size 10x14; Text '5'
   TextField "Text field_A1_0" at 172,205 size 21x14; Text '0mA'
   Bar "Bar_A1" at 192,118 size 37x97; MinimumValue 0; MaximumValue 20
      ProcessValue <- "DB001-PLC_I/O_Outputs_rAQ0.1_Scaled"

screen "03-Inputs2" 480x272, template "Main_Template"
   on GenerateScreen: SetTag("ScreenNumber", 3)
   TextField "TextField_ScreenName" at 85,46 size 309x30; Text 'PLC DIGITAL INPUTS - 2of3'
   TextField "TextField_BankLetter" at 412,50 size 62x23; Text 'BANK B'
   Group "Group_DI1.0" at 73,81 size 62x63
   Group "Group_DI1.1" at 209,81 size 62x63
   Group "Group_DI1.2" at 345,81 size 62x63
   Group "Group_DI1.3" at 73,152 size 62x63
   Group "Group_DI1.4" at 209,152 size 62x64
   Group "Group_DI1.5" at 345,152 size 62x64
   TextField "Text field_DI1.0" at 83,81 size 42x19; Text 'DI 1.0'
   Circle "Circle_DI1.0" at 86,103 size 36x36
      Appearance <- "DB001-PLC_I/O_Inputs_xDI1.0"
   TextField "Text field_DI1.1" at 219,81 size 42x19; Text 'DI 1.1'
   Circle "Circle_DI1.1" at 222,103 size 36x36
      Appearance <- "DB001-PLC_I/O_Inputs_xDI1.1"
   TextField "Text field_DI1.2" at 355,81 size 42x19; Text 'DI 1.2'
   Circle "Circle_DI1.2" at 358,103 size 36x36
      Appearance <- "DB001-PLC_I/O_Inputs_xDI1.2"
   TextField "Text field_DI1.3" at 83,152 size 42x19; Text 'DI 1.3'
   Circle "Circle_DI1.3" at 86,174 size 36x36
      Appearance <- "DB001-PLC_I/O_Inputs_xDI1.3"
   TextField "Text field_DI1.4" at 219,152 size 42x19; Text 'DI 1.4'
   Circle "Circle_DI1.4" at 222,174 size 36x36
      Appearance <- "DB001-PLC_I/O_Inputs_xDI1.4"
   TextField "Text field_DI1.5" at 355,152 size 42x19; Text 'DI 1.5'
   Circle "Circle_DI1.5" at 358,174 size 36x36
      Appearance <- "DB001-PLC_I/O_Inputs_xDI1.5"
   Button "Button_Back_1" at 411,176 size 65x40; TextOff 'BACK'
      on Press: function_efd93a16()
   Button "Button_Next" at 384,227 size 92x40; TextOff 'NEXT'
      on Press: ActivateScreen("04-Inputs3", 0)

screen "06-Outputs2" 480x272, template "Main_Template"
   on GenerateScreen: SetTag("ScreenNumber", 6)
   TextField "TextField_ScreenName" at 76,46 size 328x30; Text 'PLC DIGITAL OUTPUTS - 2of3'
   TextField "TextField_BankLetter" at 412,50 size 62x23; Text 'BANK B'
   Rectangle "Rectangle_DQ1.0" at 119,114 size 97x62
      Appearance <- "DB001-PLC_I/O_Outputs_xDQ1.0"
   TextField "Text field_DQ1.0" at 145,114 size 46x19; Text 'DQ 1.0'
   Button "Button_DQ1.0" at 131,136 size 73x32; TextOff 'Text'; TextList "ON/OFF"
      on Press: InvertBit("DB001-PLC_I/O_Outputs_xDQ1.0")
      ProcessValue <- "DB001-PLC_I/O_Outputs_xDQ0.0"
   Group "Group_DQ1.0" at 119,114 size 97x62; TextList "ON/OFF"
   Group "Group_DQ1.1" at 264,114 size 97x62; TextList "ON/OFF"
   Rectangle "Rectangle_DQ1.1" at 264,114 size 97x62
      Appearance <- "DB001-PLC_I/O_Outputs_xDQ1.1"
   TextField "Text field_DQ1.1" at 290,114 size 46x19; Text 'DQ 1.1'
   Button "Button_DQ1.1" at 276,136 size 73x32; TextOff 'Text'; TextList "ON/OFF"
      on Press: InvertBit("DB001-PLC_I/O_Outputs_xDQ1.1")
      ProcessValue <- "DB001-PLC_I/O_Outputs_xDQ0.1"
   Button "Button_Next" at 384,227 size 92x40; TextOff 'NEXT'
      on Press: ActivateScreen("07-Outputs3", 0)
   Button "Button_Back" at 384,181 size 92x40; TextOff 'BACK'
      on Press: function_efd93a16()

Template "Main_Template" 480x272
   GraphicView "Template_Background" at 0,0 size 480x272; Picture "HMI_Background"
   Button "Template_Button5_Blank" at 384,227 size 92x40; TextOff 'BLANK'
   Button "Template_Button1_Home" at 4,227 size 92x40; TextOff 'HOME'
      on Press: ActivateScreen("01-Home", 0)
   Button "Template_Button2_Inputs" at 99,227 size 92x40; TextOff 'INPUTS'
      on Press: ActivateScreen("02-Inputs1", 0)
   Button "Template_Button3_Outputs" at 194,227 size 92x40; TextOff 'OUTPUTS'
      on Press: ActivateScreen("05-Outputs1", 0)
   Button "Template_Button4_AnalogIO" at 289,227 size 92x40; TextOff 'ANALOG I/O'
      on Press: ActivateScreen("08-AnalogI/O", 0)
   IOField "Template_I/O field_Date" at 289,14 size 74x20; FormatPattern ????????
      ProcessValue <- "DB002-DateTime_sCustomDate_DDMMYY"
   IOField "Template_I/O field_Time" at 365,14 size 50x20; FormatPattern ?????
      ProcessValue <- "DB002-DateTime_sCustomTime_HHMM"
   GraphicView "TVET_Logo" at 8,2 size 220x44; Picture "TVET_Logo"

screen "07-Outputs3" 480x272, template "Main_Template"
   on GenerateScreen: SetTag("ScreenNumber", 7)
   TextField "TextField_ScreenName" at 78,46 size 325x30; Text 'PLC IO-LINK OUTPUTS - 3of3'
   TextField "Text field_Active_Input" at 24,118 size 100x17; Text 'ACTIVE - OUTPUT'
   TextField "Text field_Active_Output" at 24,140 size 89x17; Text 'ACTIVE - INPUT'
   TextField "Text field_Port_Disabled" at 24,162 size 92x17; Text 'PORT DISABLED'
   Button "Button_Back" at 384,227 size 92x40; TextOff 'BACK'
      on Press: function_efd93a16()
   TextField "Text field_X01" at 168,81 size 28x19; Text 'X01'
   Group "Group_X01" at 152,81 size 62x63
   Group "Group_X02" at 268,81 size 62x63
   Group "Group_X03" at 152,152 size 62x63
   Group "Group_X04" at 268,152 size 62x63
   TextField "Text field_X02" at 284,81 size 28x19; Text 'X02'
   TextField "Text field_X03" at 168,152 size 28x19; Text 'X03'
   TextField "Text field_X04" at 284,152 size 28x19; Text 'X04'

screen "04-Inputs3" 480x272, template "Main_Template"
   on GenerateScreen: SetTag("ScreenNumber", 4)
   Button "Button_Back" at 384,227 size 92x40; TextOff 'BACK'
      on Press: function_efd93a16()
   TextField "TextField_ScreenName" at 87,46 size 306x30; Text 'PLC IO-LINK INPUTS - 3of3'
   TextField "Text field_Active_Output" at 24,129 size 100x17; Text 'ACTIVE - OUTPUT'
   TextField "Text field_Port_Disabled" at 24,151 size 92x17; Text 'PORT DISABLED'
   Bar "Bar_X01_Temp" at 136,82 size 70x133; Unit °C; MinimumValue 0; MaximumValue 50
      ProcessValue <- "DB003-IOLink_Data_TempSensor_Data_rDeg_C"
   Group "Group_X01" at 223,81 size 82x63
   Group "Group_X02" at 325,81 size 62x63
   Group "Group_X03" at 233,152 size 62x63
   Group "Group_X04" at 325,152 size 62x63
   TextField "Text field_X01" at 250,81 size 28x19; Text 'X01'
   IOField "I/O field_X01_degC" at 229,99 size 70x20; FormatPattern s99.99; Unit  °C
      ProcessValue <- "DB003-IOLink_Data_TempSensor_Data_rDeg_C"
   IOField "I/O field_X01_degF" at 229,121 size 70x20; FormatPattern s99.99; Unit  °F
      ProcessValue <- "DB003-IOLink_Data_TempSensor_Data_rDeg_F"
   TextField "Text field_X02" at 341,81 size 28x19; Text 'X02'
   TextField "Text field_X03" at 249,152 size 28x19; Text 'X03'
   TextField "Text field_X04" at 341,152 size 28x19; Text 'X04'
*)